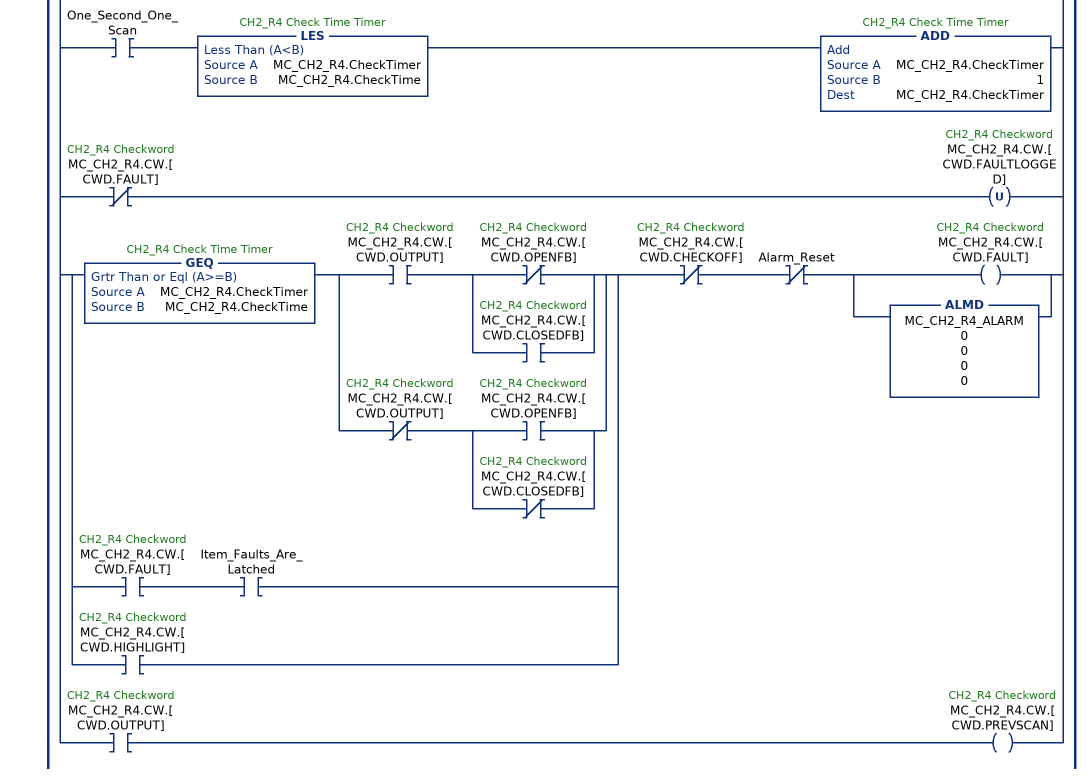
   23: [NEQ(MC_CH2_R4.DriveBits,0) OTE(MC_CH2_R4.CW.[CWD.AUTODRV]) ,[XIC(MC_CH2_R4.CW.[CWD.AUTODRV]) XIO(MC_CH2_R4.CW.[CWD.MANUAL]) ,XIC(MC_CH2_R4.CW.[CWD.MANDRV]) XIC(MC_CH2_R4.CW.[CWD.MANUAL]) ] OTE(MC_CH2_R4.CW.[CWD.OUTPUT]) ,XIC(MC_CH2_R4.CW.[CWD.OUTPUT]) OTE(MC_CH2_R4_DR) ,XIC(S:FS) [OTU(MC_CH2_R4.CW.[CWD.MANUAL]) ,LEQ(MC_CH2_R4.CheckTime,0) MOV(Default_Check_Time,MC_CH2_R4.CheckTime) ] ,[[XIC(MC_CH2_R4_O) XIO(Item_Simulation_Flag) ,XIC(Item_Simulation_Flag) XIC(MC_CH2_R4.CW.[CWD.OUTPUT]) XIO(MC_CH2_R4.CW.[CWD.SIMFAIL]) ] OTE(MC_CH2_R4.CW.[CWD.OPENFB]) ,[XIC(MC_CH2_R4_C) XIO(Item_Simulation_Flag) ,XIC(Item_Simulation_Flag) XIO(MC_CH2_R4.CW.[CWD.OUTPUT]) XIO(MC_CH2_R4.CW.[CWD.SIMFAIL]) ] OTE(MC_CH2_R4.CW.[CWD.CLOSEDFB]) ] ,[XIC(MC_CH2_R4.CW.[CWD.OUTPUT]) XIO(MC_CH2_R4.CW.[CWD.PREVSCAN]) ,XIO(MC_CH2_R4.CW.[CWD.OUTPUT]) XIC(MC_CH2_R4.CW.[CWD.PREVSCAN]) ] CLR(MC_CH2_R4.CheckTimer) ,XIC(One_Second_One_Scan) LES(MC_CH2_R4.CheckTimer,MC_CH2_R4.CheckTime) ADD(MC_CH2_R4.CheckTimer,1,MC_CH2_R4.CheckTimer) ,XIO(MC_CH2_R4.CW.[CWD.FAULT]) OTU(MC_CH2_R4.CW.[CWD.FAULTLOGGED]) ,[GEQ(MC_CH2_R4.CheckTimer,MC_CH2_R4.CheckTime) [XIC(MC_CH2_R4.CW.[CWD.OUTPUT]) [XIO(MC_CH2_R4.CW.[CWD.OPENFB]) ,XIC(MC_CH2_R4.CW.[CWD.CLOSEDFB]) ] ,XIO(MC_CH2_R4.CW.[CWD.OUTPUT]) [XIC(MC_CH2_R4.CW.[CWD.OPENFB]) ,XIO(MC_CH2_R4.CW.[CWD.CLOSEDFB]) ] ] ,XIC(MC_CH2_R4.CW.[CWD.FAULT]) XIC(Item_Faults_Are_Latched) ,XIC(MC_CH2_R4.CW.[CWD.HIGHLIGHT]) ] XIO(MC_CH2_R4.CW.[CWD.CHECKOFF]) XIO(Alarm_Reset) [OTE(MC_CH2_R4.CW.[CWD.FAULT]) ,ALMD(MC_CH2_R4_ALARM,0,0,0,0) ] ,XIC(MC_CH2_R4.CW.[CWD.OUTPUT]) OTE(MC_CH2_R4.CW.[CWD.PREVSCAN]) ];
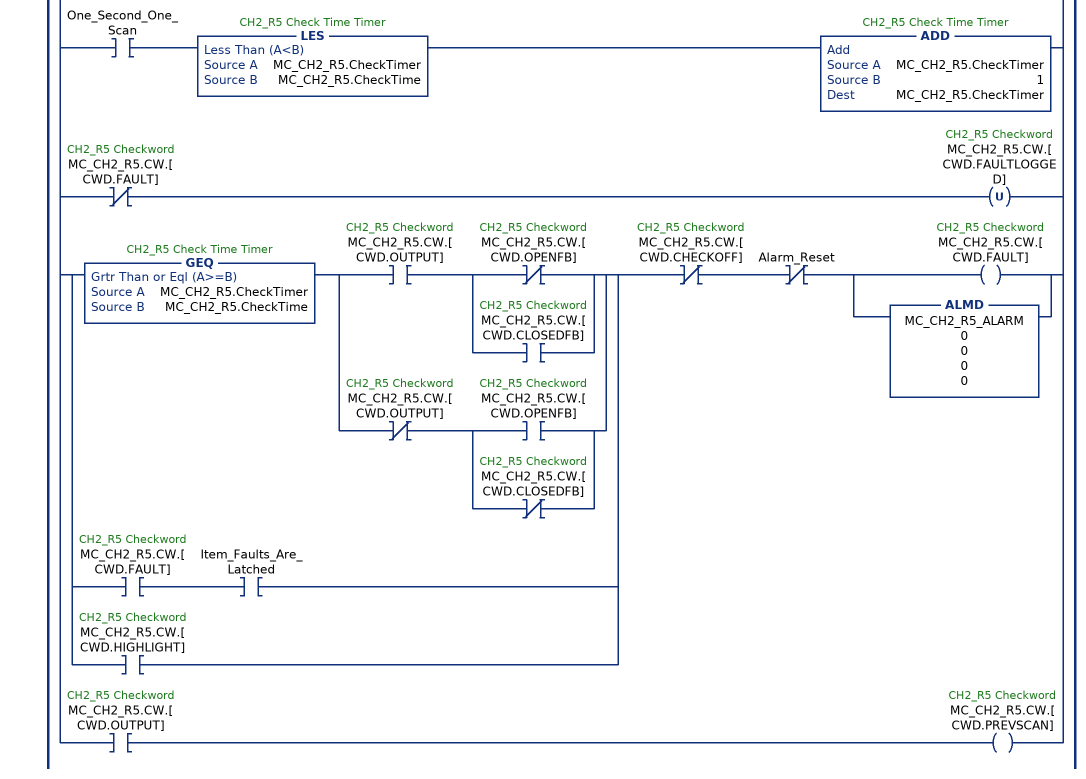
   24: [NEQ(MC_CH2_R5.DriveBits,0) OTE(MC_CH2_R5.CW.[CWD.AUTODRV]) ,[XIC(MC_CH2_R5.CW.[CWD.AUTODRV]) XIO(MC_CH2_R5.CW.[CWD.MANUAL]) ,XIC(MC_CH2_R5.CW.[CWD.MANDRV]) XIC(MC_CH2_R5.CW.[CWD.MANUAL]) ] OTE(MC_CH2_R5.CW.[CWD.OUTPUT]) ,XIC(MC_CH2_R5.CW.[CWD.OUTPUT]) OTE(MC_CH2_R5_DR) ,XIC(S:FS) [OTU(MC_CH2_R5.CW.[CWD.MANUAL]) ,LEQ(MC_CH2_R5.CheckTime,0) MOV(Default_Check_Time,MC_CH2_R5.CheckTime) ] ,[[XIC(MC_CH2_R5_O) XIO(Item_Simulation_Flag) ,XIC(Item_Simulation_Flag) XIC(MC_CH2_R5.CW.[CWD.OUTPUT]) XIO(MC_CH2_R5.CW.[CWD.SIMFAIL]) ] OTE(MC_CH2_R5.CW.[CWD.OPENFB]) ,[XIC(MC_CH2_R5_C) XIO(Item_Simulation_Flag) ,XIC(Item_Simulation_Flag) XIO(MC_CH2_R5.CW.[CWD.OUTPUT]) XIO(MC_CH2_R5.CW.[CWD.SIMFAIL]) ] OTE(MC_CH2_R5.CW.[CWD.CLOSEDFB]) ] ,[XIC(MC_CH2_R5.CW.[CWD.OUTPUT]) XIO(MC_CH2_R5.CW.[CWD.PREVSCAN]) ,XIO(MC_CH2_R5.CW.[CWD.OUTPUT]) XIC(MC_CH2_R5.CW.[CWD.PREVSCAN]) ] CLR(MC_CH2_R5.CheckTimer) ,XIC(One_Second_One_Scan) LES(MC_CH2_R5.CheckTimer,MC_CH2_R5.CheckTime) ADD(MC_CH2_R5.CheckTimer,1,MC_CH2_R5.CheckTimer) ,XIO(MC_CH2_R5.CW.[CWD.FAULT]) OTU(MC_CH2_R5.CW.[CWD.FAULTLOGGED]) ,[GEQ(MC_CH2_R5.CheckTimer,MC_CH2_R5.CheckTime) [XIC(MC_CH2_R5.CW.[CWD.OUTPUT]) [XIO(MC_CH2_R5.CW.[CWD.OPENFB]) ,XIC(MC_CH2_R5.CW.[CWD.CLOSEDFB]) ] ,XIO(MC_CH2_R5.CW.[CWD.OUTPUT]) [XIC(MC_CH2_R5.CW.[CWD.OPENFB]) ,XIO(MC_CH2_R5.CW.[CWD.CLOSEDFB]) ] ] ,XIC(MC_CH2_R5.CW.[CWD.FAULT]) XIC(Item_Faults_Are_Latched) ,XIC(MC_CH2_R5.CW.[CWD.HIGHLIGHT]) ] XIO(MC_CH2_R5.CW.[CWD.CHECKOFF]) XIO(Alarm_Reset) [OTE(MC_CH2_R5.CW.[CWD.FAULT]) ,ALMD(MC_CH2_R5_ALARM,0,0,0,0) ] ,XIC(MC_CH2_R5.CW.[CWD.OUTPUT]) OTE(MC_CH2_R5.CW.[CWD.PREVSCAN]) ];
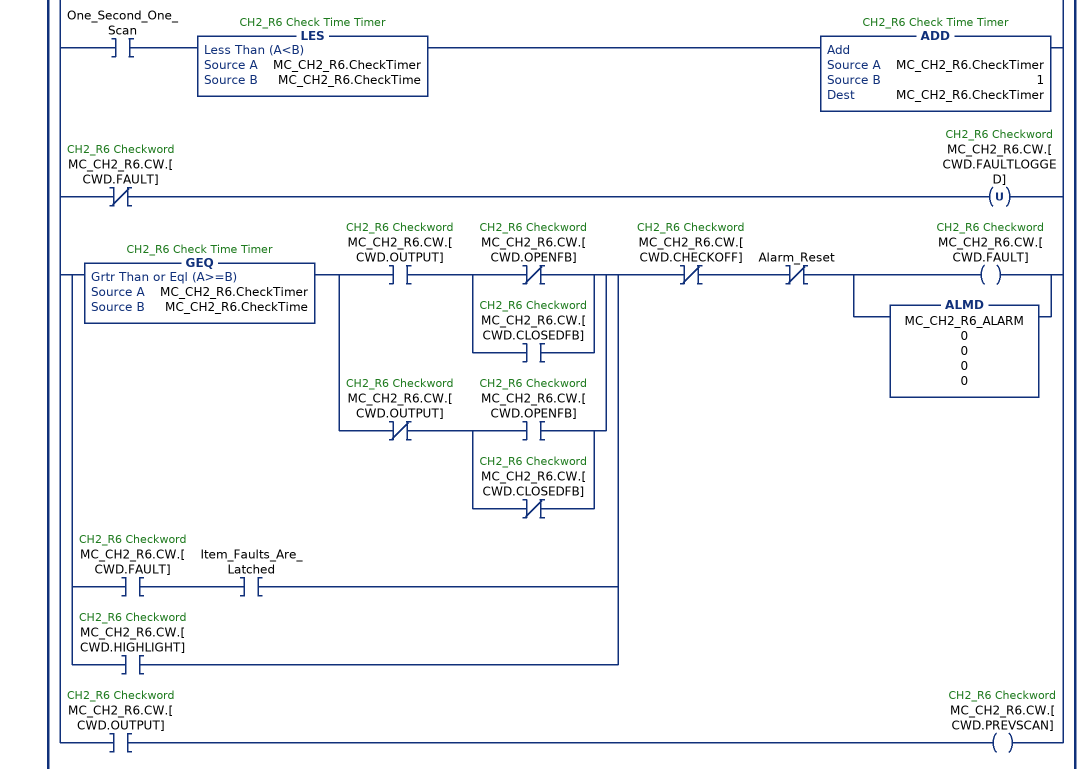
   25: [NEQ(MC_CH2_R6.DriveBits,0) OTE(MC_CH2_R6.CW.[CWD.AUTODRV]) ,[XIC(MC_CH2_R6.CW.[CWD.AUTODRV]) XIO(MC_CH2_R6.CW.[CWD.MANUAL]) ,XIC(MC_CH2_R6.CW.[CWD.MANDRV]) XIC(MC_CH2_R6.CW.[CWD.MANUAL]) ] OTE(MC_CH2_R6.CW.[CWD.OUTPUT]) ,XIC(MC_CH2_R6.CW.[CWD.OUTPUT]) OTE(MC_CH2_R6_DR) ,XIC(S:FS) [OTU(MC_CH2_R6.CW.[CWD.MANUAL]) ,LEQ(MC_CH2_R6.CheckTime,0) MOV(Default_Check_Time,MC_CH2_R6.CheckTime) ] ,[[XIC(MC_CH2_R6_O) XIO(Item_Simulation_Flag) ,XIC(Item_Simulation_Flag) XIC(MC_CH2_R6.CW.[CWD.OUTPUT]) XIO(MC_CH2_R6.CW.[CWD.SIMFAIL]) ] OTE(MC_CH2_R6.CW.[CWD.OPENFB]) ,[XIC(MC_CH2_R6_C) XIO(Item_Simulation_Flag) ,XIC(Item_Simulation_Flag) XIO(MC_CH2_R6.CW.[CWD.OUTPUT]) XIO(MC_CH2_R6.CW.[CWD.SIMFAIL]) ] OTE(MC_CH2_R6.CW.[CWD.CLOSEDFB]) ] ,[XIC(MC_CH2_R6.CW.[CWD.OUTPUT]) XIO(MC_CH2_R6.CW.[CWD.PREVSCAN]) ,XIO(MC_CH2_R6.CW.[CWD.OUTPUT]) XIC(MC_CH2_R6.CW.[CWD.PREVSCAN]) ] CLR(MC_CH2_R6.CheckTimer) ,XIC(One_Second_One_Scan) LES(MC_CH2_R6.CheckTimer,MC_CH2_R6.CheckTime) ADD(MC_CH2_R6.CheckTimer,1,MC_CH2_R6.CheckTimer) ,XIO(MC_CH2_R6.CW.[CWD.FAULT]) OTU(MC_CH2_R6.CW.[CWD.FAULTLOGGED]) ,[GEQ(MC_CH2_R6.CheckTimer,MC_CH2_R6.CheckTime) [XIC(MC_CH2_R6.CW.[CWD.OUTPUT]) [XIO(MC_CH2_R6.CW.[CWD.OPENFB]) ,XIC(MC_CH2_R6.CW.[CWD.CLOSEDFB]) ] ,XIO(MC_CH2_R6.CW.[CWD.OUTPUT]) [XIC(MC_CH2_R6.CW.[CWD.OPENFB]) ,XIO(MC_CH2_R6.CW.[CWD.CLOSEDFB]) ] ] ,XIC(MC_CH2_R6.CW.[CWD.FAULT]) XIC(Item_Faults_Are_Latched) ,XIC(MC_CH2_R6.CW.[CWD.HIGHLIGHT]) ] XIO(MC_CH2_R6.CW.[CWD.CHECKOFF]) XIO(Alarm_Reset) [OTE(MC_CH2_R6.CW.[CWD.FAULT]) ,ALMD(MC_CH2_R6_ALARM,0,0,0,0) ] ,XIC(MC_CH2_R6.CW.[CWD.OUTPUT]) OTE(MC_CH2_R6.CW.[CWD.PREVSCAN]) ];
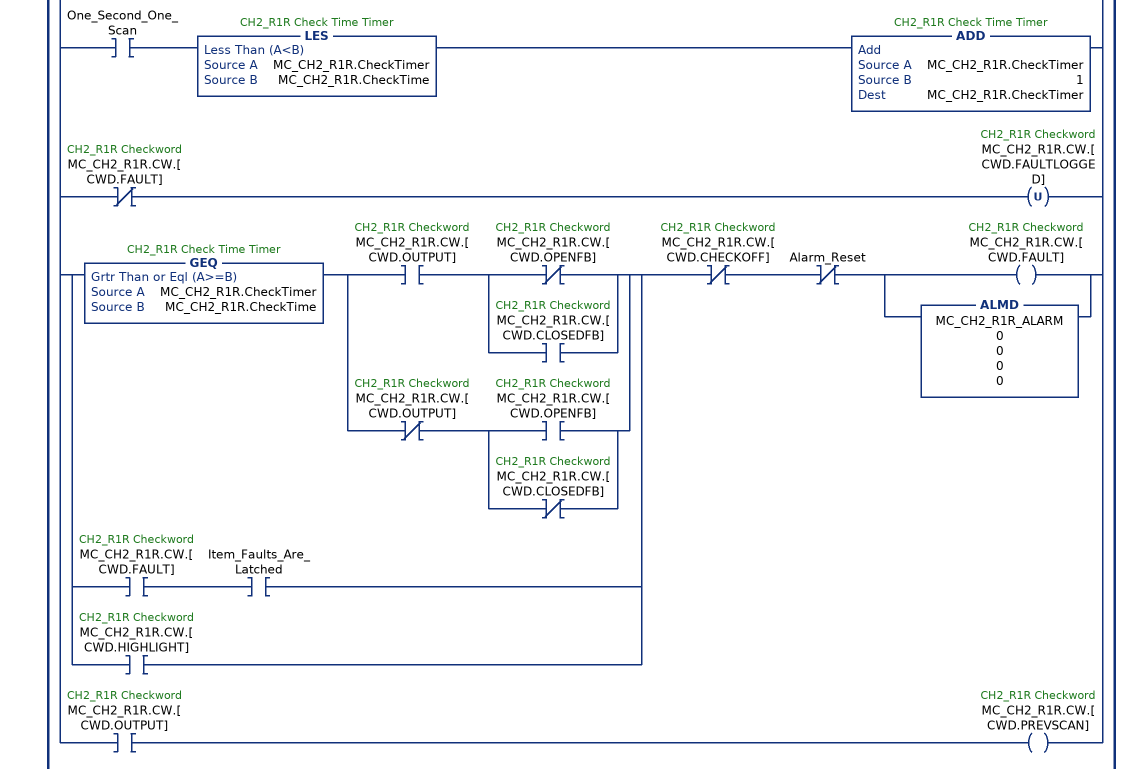
   26: [NEQ(MC_CH2_R1R.DriveBits,0) OTE(MC_CH2_R1R.CW.[CWD.AUTODRV]) ,[XIC(MC_CH2_R1R.CW.[CWD.AUTODRV]) XIO(MC_CH2_R1R.CW.[CWD.MANUAL]) ,XIC(MC_CH2_R1R.CW.[CWD.MANDRV]) XIC(MC_CH2_R1R.CW.[CWD.MANUAL]) ] OTE(MC_CH2_R1R.CW.[CWD.OUTPUT]) ,XIC(MC_CH2_R1R.CW.[CWD.OUTPUT]) OTE(MC_CH2_R1R_DR) ,XIC(S:FS) [OTU(MC_CH2_R1R.CW.[CWD.MANUAL]) ,LEQ(MC_CH2_R1R.CheckTime,0) MOV(Default_Check_Time,MC_CH2_R1R.CheckTime) ] ,[[XIC(MC_CH2_R1R_O) XIO(Item_Simulation_Flag) ,XIC(Item_Simulation_Flag) XIC(MC_CH2_R1R.CW.[CWD.OUTPUT]) XIO(MC_CH2_R1R.CW.[CWD.SIMFAIL]) ] OTE(MC_CH2_R1R.CW.[CWD.OPENFB]) ,[XIC(MC_CH2_R1R_C) XIO(Item_Simulation_Flag) ,XIC(Item_Simulation_Flag) XIO(MC_CH2_R1R.CW.[CWD.OUTPUT]) XIO(MC_CH2_R1R.CW.[CWD.SIMFAIL]) ] OTE(MC_CH2_R1R.CW.[CWD.CLOSEDFB]) ] ,[XIC(MC_CH2_R1R.CW.[CWD.OUTPUT]) XIO(MC_CH2_R1R.CW.[CWD.PREVSCAN]) ,XIO(MC_CH2_R1R.CW.[CWD.OUTPUT]) XIC(MC_CH2_R1R.CW.[CWD.PREVSCAN]) ] CLR(MC_CH2_R1R.CheckTimer) ,XIC(One_Second_One_Scan) LES(MC_CH2_R1R.CheckTimer,MC_CH2_R1R.CheckTime) ADD(MC_CH2_R1R.CheckTimer,1,MC_CH2_R1R.CheckTimer) ,XIO(MC_CH2_R1R.CW.[CWD.FAULT]) OTU(MC_CH2_R1R.CW.[CWD.FAULTLOGGED]) ,[GEQ(MC_CH2_R1R.CheckTimer,MC_CH2_R1R.CheckTime) [XIC(MC_CH2_R1R.CW.[CWD.OUTPUT]) [XIO(MC_CH2_R1R.CW.[CWD.OPENFB]) ,XIC(MC_CH2_R1R.CW.[CWD.CLOSEDFB]) ] ,XIO(MC_CH2_R1R.CW.[CWD.OUTPUT]) [XIC(MC_CH2_R1R.CW.[CWD.OPENFB]) ,XIO(MC_CH2_R1R.CW.[CWD.CLOSEDFB]) ] ] ,XIC(MC_CH2_R1R.CW.[CWD.FAULT]) XIC(Item_Faults_Are_Latched) ,XIC(MC_CH2_R1R.CW.[CWD.HIGHLIGHT]) ] XIO(MC_CH2_R1R.CW.[CWD.CHECKOFF]) XIO(Alarm_Reset) [OTE(MC_CH2_R1R.CW.[CWD.FAULT]) ,ALMD(MC_CH2_R1R_ALARM,0,0,0,0) ] ,XIC(MC_CH2_R1R.CW.[CWD.OUTPUT]) OTE(MC_CH2_R1R.CW.[CWD.PREVSCAN]) ];
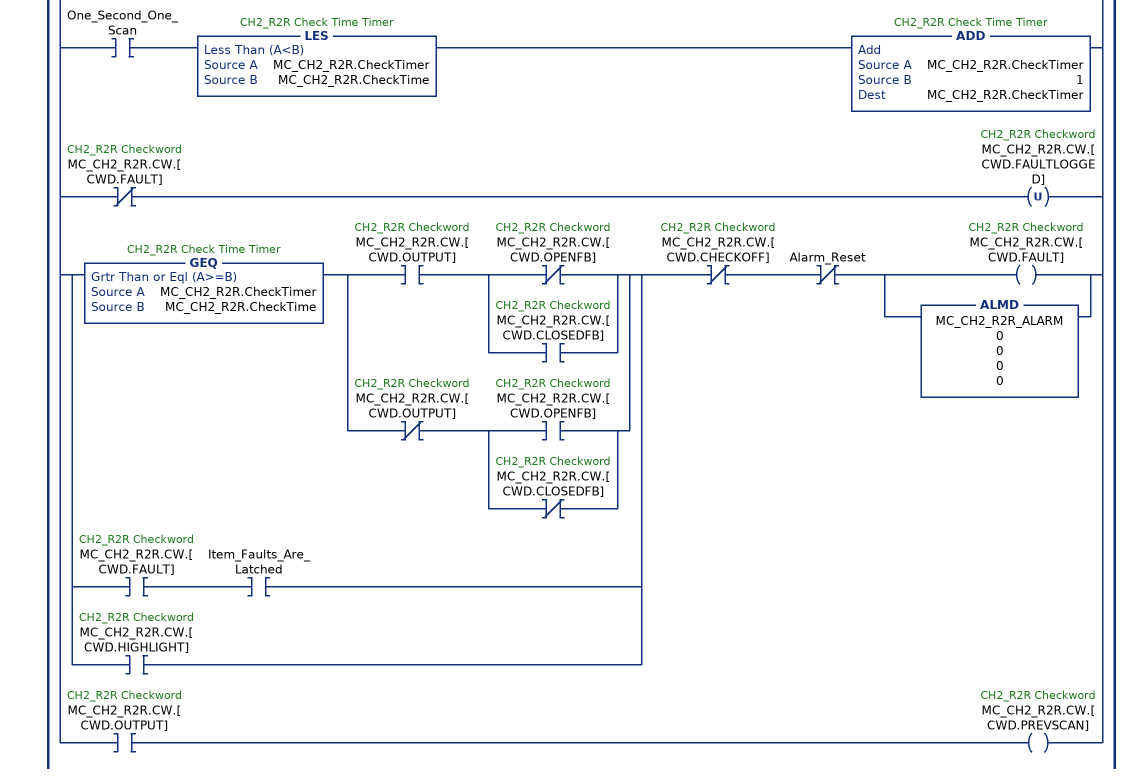
   27: [NEQ(MC_CH2_R2R.DriveBits,0) OTE(MC_CH2_R2R.CW.[CWD.AUTODRV]) ,[XIC(MC_CH2_R2R.CW.[CWD.AUTODRV]) XIO(MC_CH2_R2R.CW.[CWD.MANUAL]) ,XIC(MC_CH2_R2R.CW.[CWD.MANDRV]) XIC(MC_CH2_R2R.CW.[CWD.MANUAL]) ] OTE(MC_CH2_R2R.CW.[CWD.OUTPUT]) ,XIC(MC_CH2_R2R.CW.[CWD.OUTPUT]) OTE(MC_CH2_R2R_DR) ,XIC(S:FS) [OTU(MC_CH2_R2R.CW.[CWD.MANUAL]) ,LEQ(MC_CH2_R2R.CheckTime,0) MOV(Default_Check_Time,MC_CH2_R2R.CheckTime) ] ,[[XIC(MC_CH2_R2R_O) XIO(Item_Simulation_Flag) ,XIC(Item_Simulation_Flag) XIC(MC_CH2_R2R.CW.[CWD.OUTPUT]) XIO(MC_CH2_R2R.CW.[CWD.SIMFAIL]) ] OTE(MC_CH2_R2R.CW.[CWD.OPENFB]) ,[XIC(MC_CH2_R2R_C) XIO(Item_Simulation_Flag) ,XIC(Item_Simulation_Flag) XIO(MC_CH2_R2R.CW.[CWD.OUTPUT]) XIO(MC_CH2_R2R.CW.[CWD.SIMFAIL]) ] OTE(MC_CH2_R2R.CW.[CWD.CLOSEDFB]) ] ,[XIC(MC_CH2_R2R.CW.[CWD.OUTPUT]) XIO(MC_CH2_R2R.CW.[CWD.PREVSCAN]) ,XIO(MC_CH2_R2R.CW.[CWD.OUTPUT]) XIC(MC_CH2_R2R.CW.[CWD.PREVSCAN]) ] CLR(MC_CH2_R2R.CheckTimer) ,XIC(One_Second_One_Scan) LES(MC_CH2_R2R.CheckTimer,MC_CH2_R2R.CheckTime) ADD(MC_CH2_R2R.CheckTimer,1,MC_CH2_R2R.CheckTimer) ,XIO(MC_CH2_R2R.CW.[CWD.FAULT]) OTU(MC_CH2_R2R.CW.[CWD.FAULTLOGGED]) ,[GEQ(MC_CH2_R2R.CheckTimer,MC_CH2_R2R.CheckTime) [XIC(MC_CH2_R2R.CW.[CWD.OUTPUT]) [XIO(MC_CH2_R2R.CW.[CWD.OPENFB]) ,XIC(MC_CH2_R2R.CW.[CWD.CLOSEDFB]) ] ,XIO(MC_CH2_R2R.CW.[CWD.OUTPUT]) [XIC(MC_CH2_R2R.CW.[CWD.OPENFB]) ,XIO(MC_CH2_R2R.CW.[CWD.CLOSEDFB]) ] ] ,XIC(MC_CH2_R2R.CW.[CWD.FAULT]) XIC(Item_Faults_Are_Latched) ,XIC(MC_CH2_R2R.CW.[CWD.HIGHLIGHT]) ] XIO(MC_CH2_R2R.CW.[CWD.CHECKOFF]) XIO(Alarm_Reset) [OTE(MC_CH2_R2R.CW.[CWD.FAULT]) ,ALMD(MC_CH2_R2R_ALARM,0,0,0,0) ] ,XIC(MC_CH2_R2R.CW.[CWD.OUTPUT]) OTE(MC_CH2_R2R.CW.[CWD.PREVSCAN]) ];
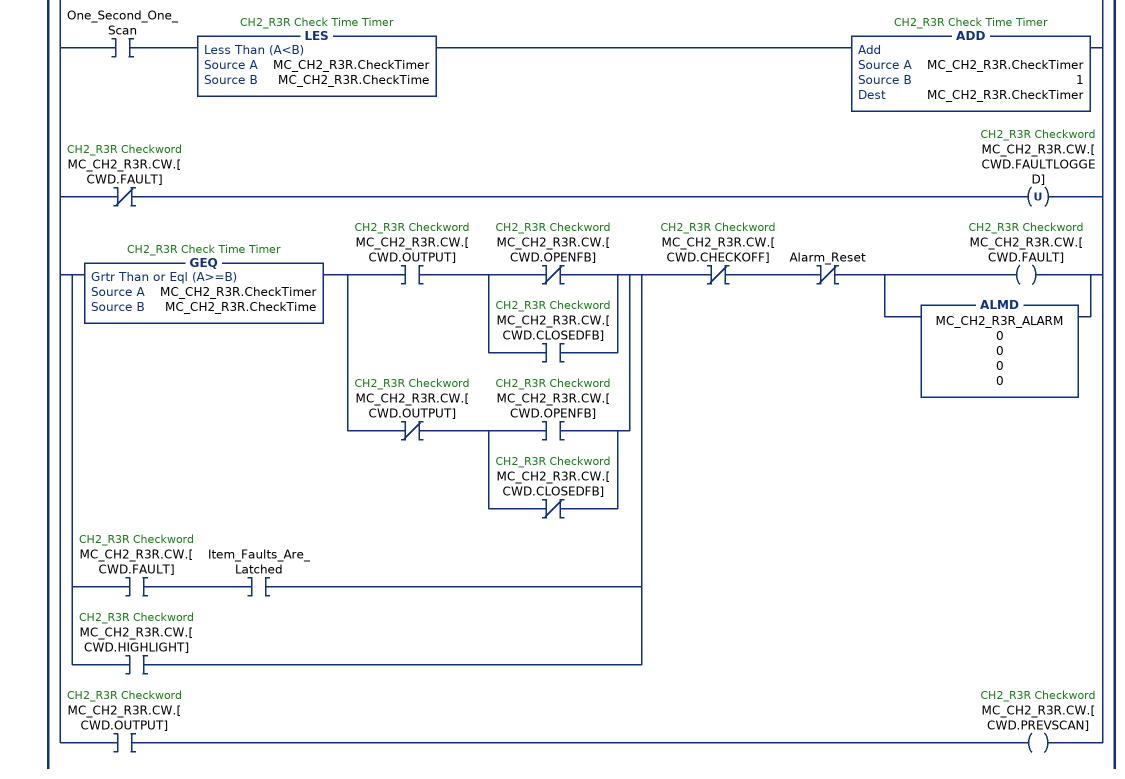
   28: [NEQ(MC_CH2_R3R.DriveBits,0) OTE(MC_CH2_R3R.CW.[CWD.AUTODRV]) ,[XIC(MC_CH2_R3R.CW.[CWD.AUTODRV]) XIO(MC_CH2_R3R.CW.[CWD.MANUAL]) ,XIC(MC_CH2_R3R.CW.[CWD.MANDRV]) XIC(MC_CH2_R3R.CW.[CWD.MANUAL]) ] OTE(MC_CH2_R3R.CW.[CWD.OUTPUT]) ,XIC(MC_CH2_R3R.CW.[CWD.OUTPUT]) OTE(MC_CH2_R3R_DR) ,XIC(S:FS) [OTU(MC_CH2_R3R.CW.[CWD.MANUAL]) ,LEQ(MC_CH2_R3R.CheckTime,0) MOV(Default_Check_Time,MC_CH2_R3R.CheckTime) ] ,[[XIC(MC_CH2_R3R_O) XIO(Item_Simulation_Flag) ,XIC(Item_Simulation_Flag) XIC(MC_CH2_R3R.CW.[CWD.OUTPUT]) XIO(MC_CH2_R3R.CW.[CWD.SIMFAIL]) ] OTE(MC_CH2_R3R.CW.[CWD.OPENFB]) ,[XIC(MC_CH2_R3R_C) XIO(Item_Simulation_Flag) ,XIC(Item_Simulation_Flag) XIO(MC_CH2_R3R.CW.[CWD.OUTPUT]) XIO(MC_CH2_R3R.CW.[CWD.SIMFAIL]) ] OTE(MC_CH2_R3R.CW.[CWD.CLOSEDFB]) ] ,[XIC(MC_CH2_R3R.CW.[CWD.OUTPUT]) XIO(MC_CH2_R3R.CW.[CWD.PREVSCAN]) ,XIO(MC_CH2_R3R.CW.[CWD.OUTPUT]) XIC(MC_CH2_R3R.CW.[CWD.PREVSCAN]) ] CLR(MC_CH2_R3R.CheckTimer) ,XIC(One_Second_One_Scan) LES(MC_CH2_R3R.CheckTimer,MC_CH2_R3R.CheckTime) ADD(MC_CH2_R3R.CheckTimer,1,MC_CH2_R3R.CheckTimer) ,XIO(MC_CH2_R3R.CW.[CWD.FAULT]) OTU(MC_CH2_R3R.CW.[CWD.FAULTLOGGED]) ,[GEQ(MC_CH2_R3R.CheckTimer,MC_CH2_R3R.CheckTime) [XIC(MC_CH2_R3R.CW.[CWD.OUTPUT]) [XIO(MC_CH2_R3R.CW.[CWD.OPENFB]) ,XIC(MC_CH2_R3R.CW.[CWD.CLOSEDFB]) ] ,XIO(MC_CH2_R3R.CW.[CWD.OUTPUT]) [XIC(MC_CH2_R3R.CW.[CWD.OPENFB]) ,XIO(MC_CH2_R3R.CW.[CWD.CLOSEDFB]) ] ] ,XIC(MC_CH2_R3R.CW.[CWD.FAULT]) XIC(Item_Faults_Are_Latched) ,XIC(MC_CH2_R3R.CW.[CWD.HIGHLIGHT]) ] XIO(MC_CH2_R3R.CW.[CWD.CHECKOFF]) XIO(Alarm_Reset) [OTE(MC_CH2_R3R.CW.[CWD.FAULT]) ,ALMD(MC_CH2_R3R_ALARM,0,0,0,0) ] ,XIC(MC_CH2_R3R.CW.[CWD.OUTPUT]) OTE(MC_CH2_R3R.CW.[CWD.PREVSCAN]) ];
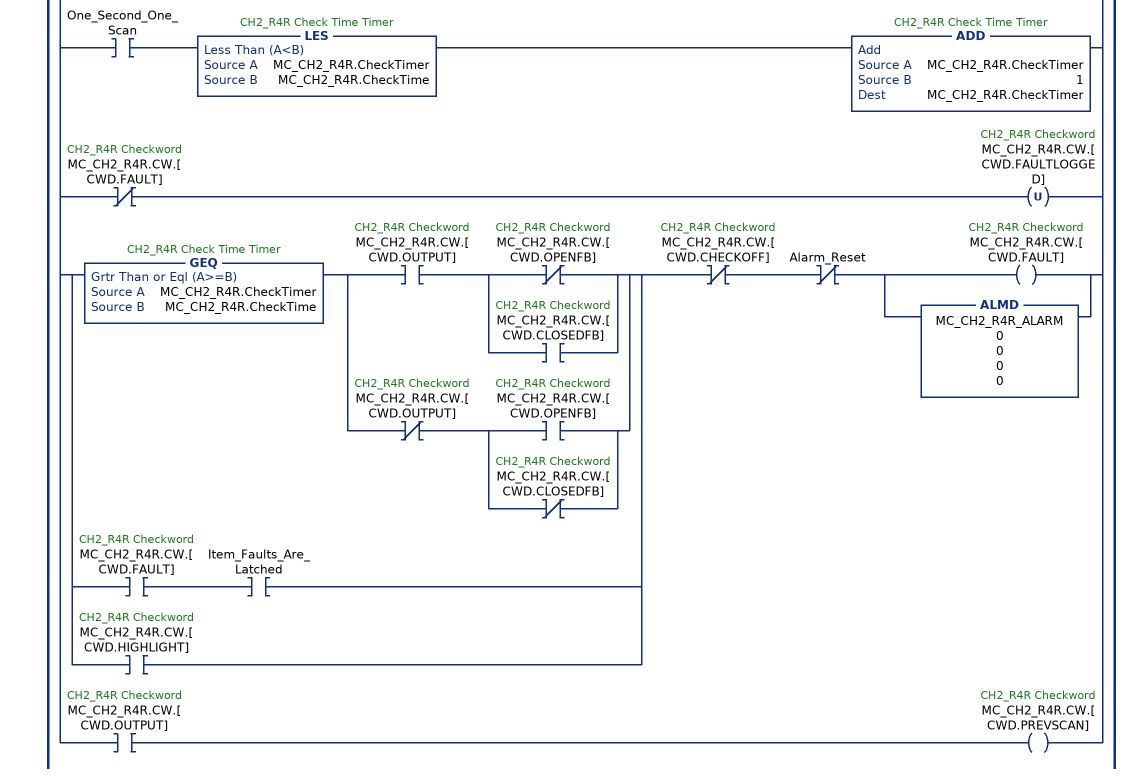
   29: [NEQ(MC_CH2_R4R.DriveBits,0) OTE(MC_CH2_R4R.CW.[CWD.AUTODRV]) ,[XIC(MC_CH2_R4R.CW.[CWD.AUTODRV]) XIO(MC_CH2_R4R.CW.[CWD.MANUAL]) ,XIC(MC_CH2_R4R.CW.[CWD.MANDRV]) XIC(MC_CH2_R4R.CW.[CWD.MANUAL]) ] OTE(MC_CH2_R4R.CW.[CWD.OUTPUT]) ,XIC(MC_CH2_R4R.CW.[CWD.OUTPUT]) OTE(MC_CH2_R4R_DR) ,XIC(S:FS) [OTU(MC_CH2_R4R.CW.[CWD.MANUAL]) ,LEQ(MC_CH2_R4R.CheckTime,0) MOV(Default_Check_Time,MC_CH2_R4R.CheckTime) ] ,[[XIC(MC_CH2_R4R_O) XIO(Item_Simulation_Flag) ,XIC(Item_Simulation_Flag) XIC(MC_CH2_R4R.CW.[CWD.OUTPUT]) XIO(MC_CH2_R4R.CW.[CWD.SIMFAIL]) ] OTE(MC_CH2_R4R.CW.[CWD.OPENFB]) ,[XIC(MC_CH2_R4R_C) XIO(Item_Simulation_Flag) ,XIC(Item_Simulation_Flag) XIO(MC_CH2_R4R.CW.[CWD.OUTPUT]) XIO(MC_CH2_R4R.CW.[CWD.SIMFAIL]) ] OTE(MC_CH2_R4R.CW.[CWD.CLOSEDFB]) ] ,[XIC(MC_CH2_R4R.CW.[CWD.OUTPUT]) XIO(MC_CH2_R4R.CW.[CWD.PREVSCAN]) ,XIO(MC_CH2_R4R.CW.[CWD.OUTPUT]) XIC(MC_CH2_R4R.CW.[CWD.PREVSCAN]) ] CLR(MC_CH2_R4R.CheckTimer) ,XIC(One_Second_One_Scan) LES(MC_CH2_R4R.CheckTimer,MC_CH2_R4R.CheckTime) ADD(MC_CH2_R4R.CheckTimer,1,MC_CH2_R4R.CheckTimer) ,XIO(MC_CH2_R4R.CW.[CWD.FAULT]) OTU(MC_CH2_R4R.CW.[CWD.FAULTLOGGED]) ,[GEQ(MC_CH2_R4R.CheckTimer,MC_CH2_R4R.CheckTime) [XIC(MC_CH2_R4R.CW.[CWD.OUTPUT]) [XIO(MC_CH2_R4R.CW.[CWD.OPENFB]) ,XIC(MC_CH2_R4R.CW.[CWD.CLOSEDFB]) ] ,XIO(MC_CH2_R4R.CW.[CWD.OUTPUT]) [XIC(MC_CH2_R4R.CW.[CWD.OPENFB]) ,XIO(MC_CH2_R4R.CW.[CWD.CLOSEDFB]) ] ] ,XIC(MC_CH2_R4R.CW.[CWD.FAULT]) XIC(Item_Faults_Are_Latched) ,XIC(MC_CH2_R4R.CW.[CWD.HIGHLIGHT]) ] XIO(MC_CH2_R4R.CW.[CWD.CHECKOFF]) XIO(Alarm_Reset) [OTE(MC_CH2_R4R.CW.[CWD.FAULT]) ,ALMD(MC_CH2_R4R_ALARM,0,0,0,0) ] ,XIC(MC_CH2_R4R.CW.[CWD.OUTPUT]) OTE(MC_CH2_R4R.CW.[CWD.PREVSCAN]) ];
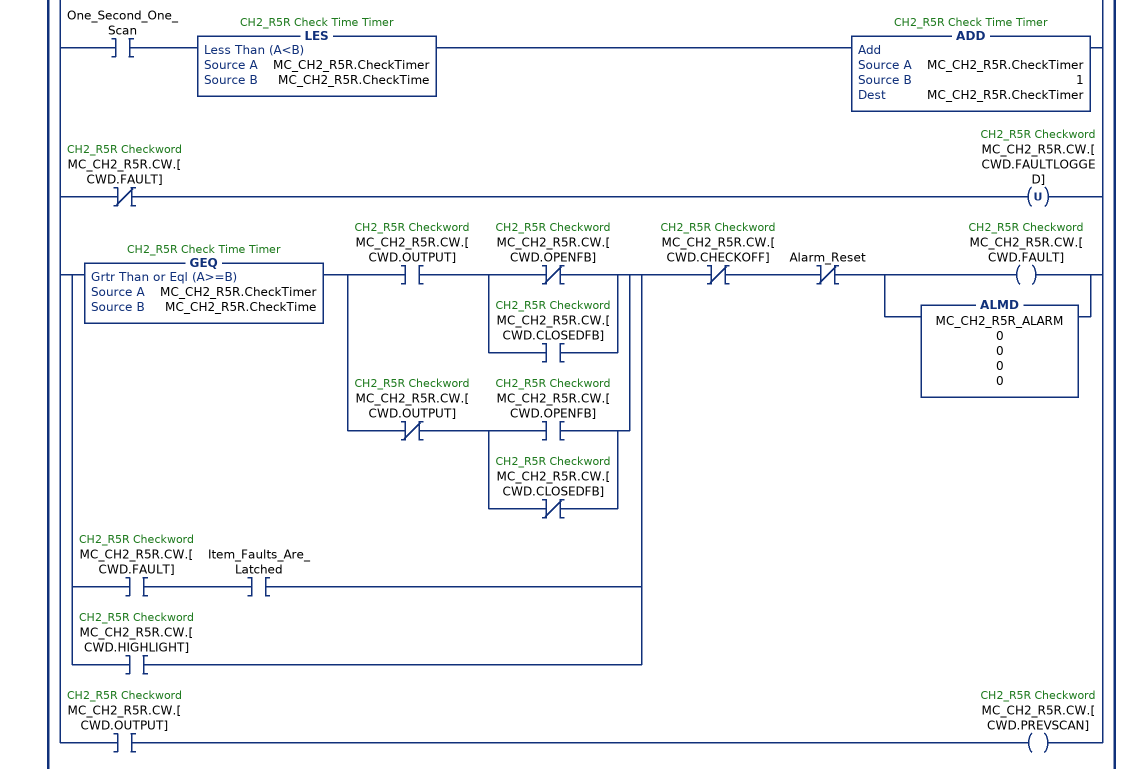
   30: [NEQ(MC_CH2_R5R.DriveBits,0) OTE(MC_CH2_R5R.CW.[CWD.AUTODRV]) ,[XIC(MC_CH2_R5R.CW.[CWD.AUTODRV]) XIO(MC_CH2_R5R.CW.[CWD.MANUAL]) ,XIC(MC_CH2_R5R.CW.[CWD.MANDRV]) XIC(MC_CH2_R5R.CW.[CWD.MANUAL]) ] OTE(MC_CH2_R5R.CW.[CWD.OUTPUT]) ,XIC(MC_CH2_R5R.CW.[CWD.OUTPUT]) OTE(MC_CH2_R5R_DR) ,XIC(S:FS) [OTU(MC_CH2_R5R.CW.[CWD.MANUAL]) ,LEQ(MC_CH2_R5R.CheckTime,0) MOV(Default_Check_Time,MC_CH2_R5R.CheckTime) ] ,[[XIC(MC_CH2_R5R_O) XIO(Item_Simulation_Flag) ,XIC(Item_Simulation_Flag) XIC(MC_CH2_R5R.CW.[CWD.OUTPUT]) XIO(MC_CH2_R5R.CW.[CWD.SIMFAIL]) ] OTE(MC_CH2_R5R.CW.[CWD.OPENFB]) ,[XIC(MC_CH2_R5R_C) XIO(Item_Simulation_Flag) ,XIC(Item_Simulation_Flag) XIO(MC_CH2_R5R.CW.[CWD.OUTPUT]) XIO(MC_CH2_R5R.CW.[CWD.SIMFAIL]) ] OTE(MC_CH2_R5R.CW.[CWD.CLOSEDFB]) ] ,[XIC(MC_CH2_R5R.CW.[CWD.OUTPUT]) XIO(MC_CH2_R5R.CW.[CWD.PREVSCAN]) ,XIO(MC_CH2_R5R.CW.[CWD.OUTPUT]) XIC(MC_CH2_R5R.CW.[CWD.PREVSCAN]) ] CLR(MC_CH2_R5R.CheckTimer) ,XIC(One_Second_One_Scan) LES(MC_CH2_R5R.CheckTimer,MC_CH2_R5R.CheckTime) ADD(MC_CH2_R5R.CheckTimer,1,MC_CH2_R5R.CheckTimer) ,XIO(MC_CH2_R5R.CW.[CWD.FAULT]) OTU(MC_CH2_R5R.CW.[CWD.FAULTLOGGED]) ,[GEQ(MC_CH2_R5R.CheckTimer,MC_CH2_R5R.CheckTime) [XIC(MC_CH2_R5R.CW.[CWD.OUTPUT]) [XIO(MC_CH2_R5R.CW.[CWD.OPENFB]) ,XIC(MC_CH2_R5R.CW.[CWD.CLOSEDFB]) ] ,XIO(MC_CH2_R5R.CW.[CWD.OUTPUT]) [XIC(MC_CH2_R5R.CW.[CWD.OPENFB]) ,XIO(MC_CH2_R5R.CW.[CWD.CLOSEDFB]) ] ] ,XIC(MC_CH2_R5R.CW.[CWD.FAULT]) XIC(Item_Faults_Are_Latched) ,XIC(MC_CH2_R5R.CW.[CWD.HIGHLIGHT]) ] XIO(MC_CH2_R5R.CW.[CWD.CHECKOFF]) XIO(Alarm_Reset) [OTE(MC_CH2_R5R.CW.[CWD.FAULT]) ,ALMD(MC_CH2_R5R_ALARM,0,0,0,0) ] ,XIC(MC_CH2_R5R.CW.[CWD.OUTPUT]) OTE(MC_CH2_R5R.CW.[CWD.PREVSCAN]) ];
